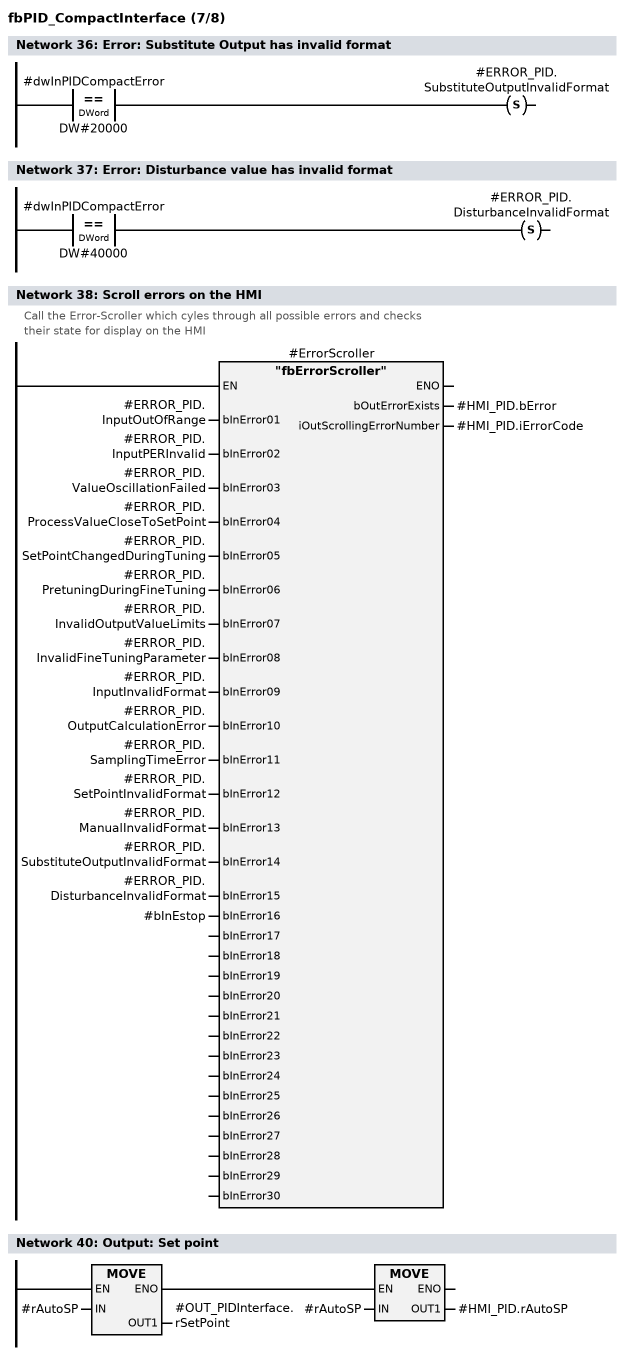
   RUNG wire#powerrail
      { S7_Templates := "SrcType := DWord" } EQ_Contact(in1 := #dwInPIDCompactError, in2 := DW#20000)
      S_Coil( #ERROR_PID.SubstituteOutputInvalidFormat )
   END_RUNG
   // the same network as SCL:
   IF #dwInPIDCompactError = DW#20000 THEN #ERROR_PID.SubstituteOutputInvalidFormat := TRUE; END_IF;
END_REGION

REGION Network 37: Error: Disturbance value has invalid format
   RUNG wire#powerrail
      { S7_Templates := "SrcType := DWord" } EQ_Contact(in1 := #dwInPIDCompactError, in2 := DW#40000)
      S_Coil( #ERROR_PID.DisturbanceInvalidFormat )
   END_RUNG
   // the same network as SCL:
   IF #dwInPIDCompactError = DW#40000 THEN #ERROR_PID.DisturbanceInvalidFormat := TRUE; END_IF;
END_REGION

REGION Network 38: Scroll errors on the HMI
   // Call the Error-Scroller which cyles through all possible errors and checks 
   // their state for display on the HMI
   RUNG wire#powerrail
      #ErrorScroller(bInError01 := #ERROR_PID.InputOutOfRange, bInError02 := #ERROR_PID.InputPERInvalid, bInError03 := #ERROR_PID.ValueOscillationFailed, bInError04 := #ERROR_PID.ProcessValueCloseToSetPoint, bInError05 := #ERROR_PID.SetPointChangedDuringTuning, bInError06 := #ERROR_PID.PretuningDuringFineTuning, bInError07 := #ERROR_PID.InvalidOutputValueLimits, bInError08 := #ERROR_PID.InvalidFineTuningParameter, bInError09 := #ERROR_PID.InputInvalidFormat, bInError10 := #ERROR_PID.OutputCalculationError, bInError11 := #ERROR_PID.SamplingTimeError, bInError12 := #ERROR_PID.SetPointInvalidFormat, bInError13 := #ERROR_PID.ManualInvalidFormat, bInError14 := #ERROR_PID.SubstituteOutputInvalidFormat, bInError15 := #ERROR_PID.DisturbanceInvalidFormat, bInError16 := #bInEstop, bInError17 :=, bInError18 :=, bInError19 :=, bInError20 :=, bInError21 :=, bInError22 :=, bInError23 :=, bInError24 :=, bInError25 :=, bInError26 :=, bInError27 :=, bInError28 :=, bInError29 :=, bInError30 :=, bOutErrorExists => #HMI_PID.bError, iOutScrollingErrorNumber => #HMI_PID.iErrorCode)
   END_RUNG
   // the same network as SCL:
   #ErrorScroller(bInError01 := #ERROR_PID.InputOutOfRange,   // "fbErrorScroller"
                  bInError02 := #ERROR_PID.InputPERInvalid,
                  bInError03 := #ERROR_PID.ValueOscillationFailed,
                  bInError04 := #ERROR_PID.ProcessValueCloseToSetPoint,
                  bInError05 := #ERROR_PID.SetPointChangedDuringTuning,
                  bInError06 := #ERROR_PID.PretuningDuringFineTuning,
                  bInError07 := #ERROR_PID.InvalidOutputValueLimits,
                  bInError08 := #ERROR_PID.InvalidFineTuningParameter,
                  bInError09 := #ERROR_PID.InputInvalidFormat,
                  bInError10 := #ERROR_PID.OutputCalculationError,
                  bInError11 := #ERROR_PID.SamplingTimeError,
                  bInError12 := #ERROR_PID.SetPointInvalidFormat,
                  bInError13 := #ERROR_PID.ManualInvalidFormat,
                  bInError14 := #ERROR_PID.SubstituteOutputInvalidFormat,
                  bInError15 := #ERROR_PID.DisturbanceInvalidFormat,
                  bInError16 := #bInEstop,
                  bOutErrorExists => #HMI_PID.bError,
                  iOutScrollingErrorNumber => #HMI_PID.iErrorCode);
END_REGION

REGION Network 39: --------------------------------------------------------- Outputs ------------------------------------------------------------------
END_REGION

REGION Network 40: Output: Set point
   RUNG wire#powerrail
      Move(in := #rAutoSP, out1 => #OUT_PIDInterface.rSetPoint)
      Move(in := #rAutoSP, out1 => #HMI_PID.rAutoSP)
   END_RUNG
   // the same network as SCL:
   #OUT_PIDInterface.rSetPoint := #rAutoSP;
   #HMI_PID.rAutoSP := #rAutoSP;
END_REGION

REGION Network 41: Output: Process value
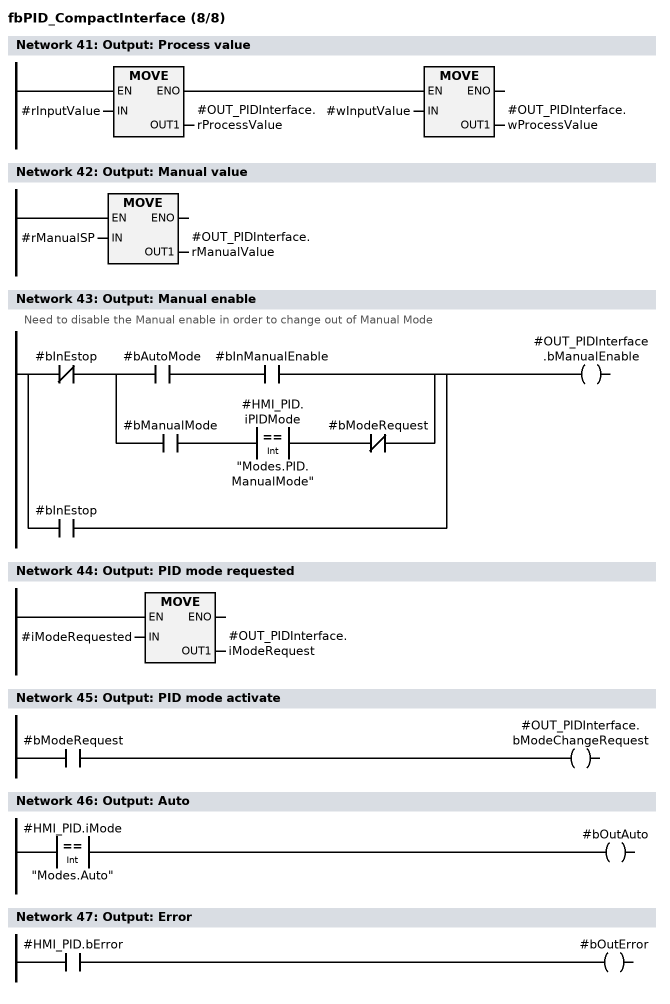
   RUNG wire#powerrail
      Move(in := #rInputValue, out1 => #OUT_PIDInterface.rProcessValue)
      Move(in := #wInputValue, out1 => #OUT_PIDInterface.wProcessValue)
   END_RUNG
   // the same network as SCL:
   #OUT_PIDInterface.rProcessValue := #rInputValue;
   #OUT_PIDInterface.wProcessValue := #wInputValue;
END_REGION

REGION Network 42: Output: Manual value
   RUNG wire#powerrail
      Move(in := #rManualSP, out1 => #OUT_PIDInterface.rManualValue)
   END_RUNG
   // the same network as SCL:
   #OUT_PIDInterface.rManualValue := #rManualSP;
END_REGION

REGION Network 43: Output: Manual enable
   // Need to disable the Manual enable in order to change out of Manual Mode
   RUNG wire#powerrail
      I_Contact( #bInEstop )
      wire#w1
      Contact( #bAutoMode )
      Contact( #bInManualEnable )
      wire#w2
      Coil( #OUT_PIDInterface.bManualEnable )
   END_RUNG
   RUNG wire#w1
      Contact( #bManualMode )
      { S7_Templates := "SrcType := Int" } EQ_Contact(in1 := #HMI_PID.iPIDMode, in2 := "Modes.PID.ManualMode")
      I_Contact( #bModeRequest )
   END_RUNG wire#w2
   RUNG wire#powerrail
      Contact( #bInEstop )
   END_RUNG wire#w2
   // the same network as SCL:
   #OUT_PIDInterface.bManualEnable := (NOT #bInEstop AND ((#bAutoMode AND #bInManualEnable) OR (#bManualMode AND (#HMI_PID.iPIDMode = "Modes.PID.ManualMode") AND NOT #bModeRequest))) OR #bInEstop;
END_REGION

REGION Network 44: Output: PID mode requested
   RUNG wire#powerrail
      Move(in := #iModeRequested, out1 => #OUT_PIDInterface.iModeRequest)
   END_RUNG
   // the same network as SCL:
   #OUT_PIDInterface.iModeRequest := #iModeRequested;
END_REGION

REGION Network 45: Output: PID mode activate
   RUNG wire#powerrail
      Contact( #bModeRequest )
      Coil( #OUT_PIDInterface.bModeChangeRequest )
   END_RUNG
   // the same network as SCL:
   #OUT_PIDInterface.bModeChangeRequest := #bModeRequest;
END_REGION

REGION Network 46: Output: Auto
   RUNG wire#powerrail
      { S7_Templates := "SrcType := Int" } EQ_Contact(in1 := #HMI_PID.iMode, in2 := "Modes.Auto")
      Coil( #bOutAuto )
   END_RUNG
   // the same network as SCL:
   #bOutAuto := #HMI_PID.iMode = "Modes.Auto";
END_REGION

REGION Network 47: Output: Error
   RUNG wire#powerrail
      Contact( #HMI_PID.bError )
      Coil( #bOutError )
   END_RUNG
   // the same network as SCL:
   #bOutError := #HMI_PID.bError;
END_REGION
END_FUNCTION_BLOCK

// folder: Library Blocks/Resources/Communication

FUNCTION_BLOCK "fbAsyncParameterRW_VFD"   // FB125, LAD
TITLE = VFD Acylic Parameter Read and Write
{ S7_Optimized_Access := 'FALSE' }
AUTHOR : JRM
NAME : VFD
VERSION : 0.1
// This block works on Siemens MicroMasters and G120 VFDs
   VAR_TEMP   // added for the SCL form of the ladder/FBD networks
      _w1 : Bool;
   END_VAR
BEGIN

REGION Network 1: ------------------------ Set Values --------------------------
END_REGION

REGION Network 2: Check valid state
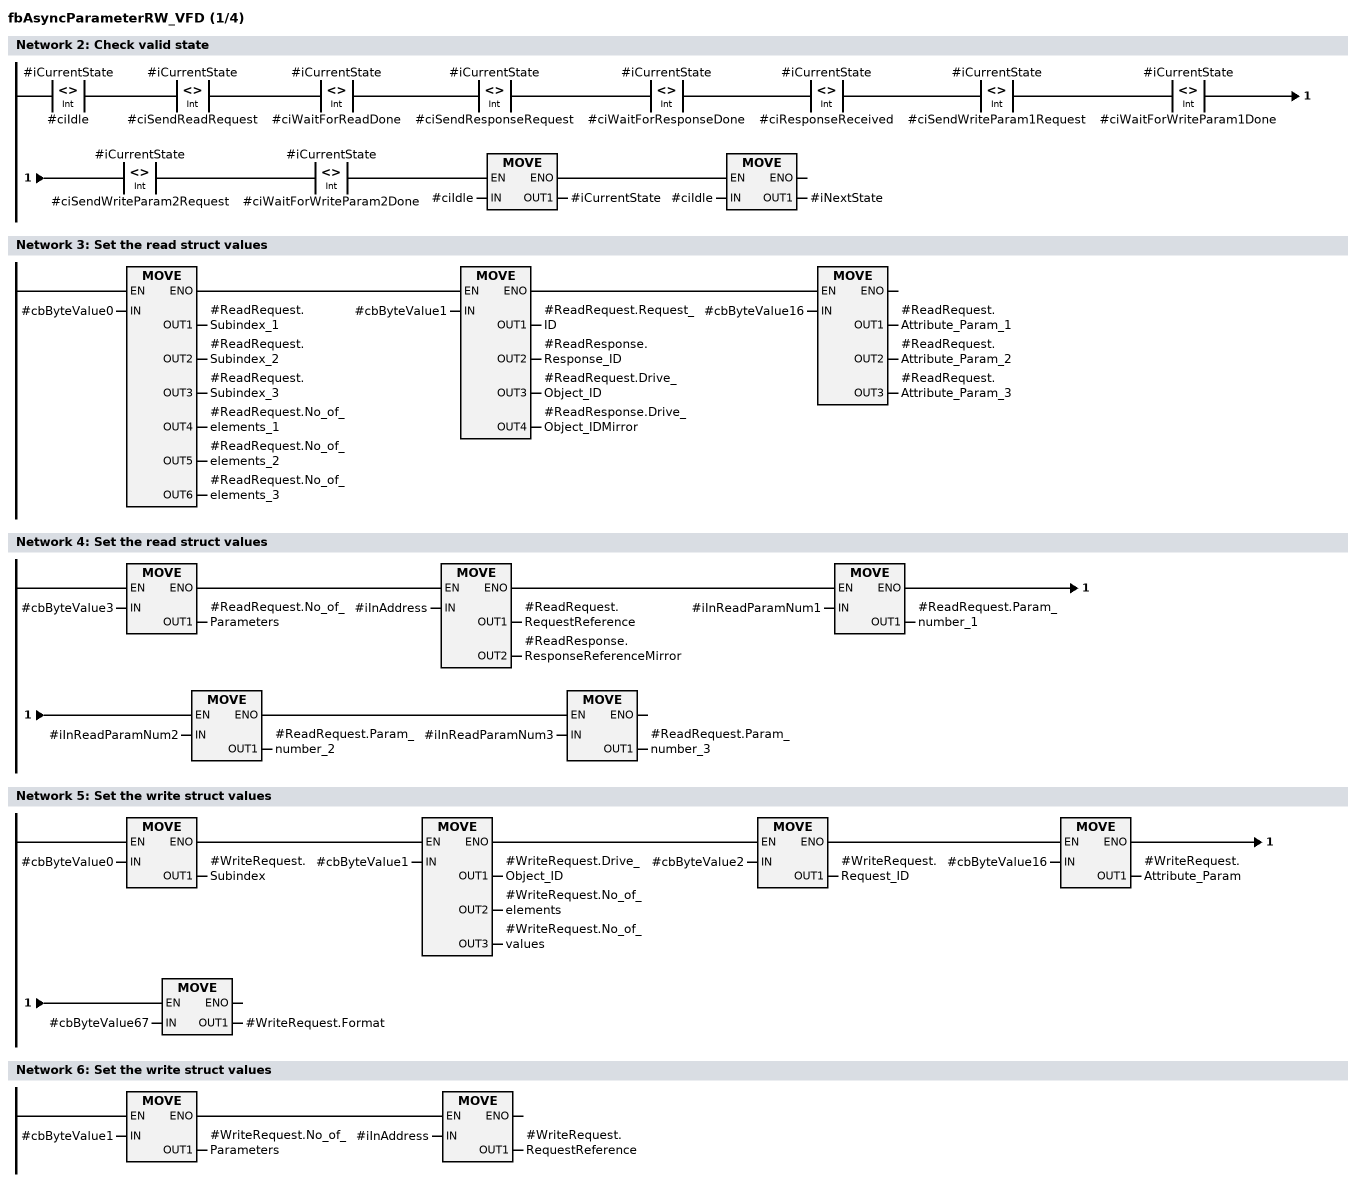
   RUNG wire#powerrail
      { S7_Templates := "SrcType := Int" } NE_Contact(in1 := #iCurrentState, in2 := #ciIdle)
      { S7_Templates := "SrcType := Int" } NE_Contact(in1 := #iCurrentState, in2 := #ciSendReadRequest)
      { S7_Templates := "SrcType := Int" } NE_Contact(in1 := #iCurrentState, in2 := #ciWaitForReadDone)
      { S7_Templates := "SrcType := Int" } NE_Contact(in1 := #iCurrentState, in2 := #ciSendResponseRequest)
      { S7_Templates := "SrcType := Int" } NE_Contact(in1 := #iCurrentState, in2 := #ciWaitForResponseDone)
      { S7_Templates := "SrcType := Int" } NE_Contact(in1 := #iCurrentState, in2 := #ciResponseReceived)
      { S7_Templates := "SrcType := Int" } NE_Contact(in1 := #iCurrentState, in2 := #ciSendWriteParam1Request)
      { S7_Templates := "SrcType := Int" } NE_Contact(in1 := #iCurrentState, in2 := #ciWaitForWriteParam1Done)
      { S7_Templates := "SrcType := Int" } NE_Contact(in1 := #iCurrentState, in2 := #ciSendWriteParam2Request)
      { S7_Templates := "SrcType := Int" } NE_Contact(in1 := #iCurrentState, in2 := #ciWaitForWriteParam2Done)
      { S7_GenerateENO := "TRUE" } Move(in := #ciIdle, out1 => #iCurrentState)
      { S7_GenerateENO := "TRUE" } Move(in := #ciIdle, out1 => #iNextState)
   END_RUNG
   // the same network as SCL:
   // ENO of a box is taken as its EN; it also drops when the box reports an error
   #_w1 := (#iCurrentState <> #ciIdle) AND (#iCurrentState <> #ciSendReadRequest) AND (#iCurrentState <> #ciWaitForReadDone) AND (#iCurrentState <> #ciSendResponseRequest) AND (#iCurrentState <> #ciWaitForResponseDone) AND (#iCurrentState <> #ciResponseReceived) AND (#iCurrentState <> #ciSendWriteParam1Request) AND (#iCurrentState <> #ciWaitForWriteParam1Done) AND (#iCurrentState <> #ciSendWriteParam2Request) AND (#iCurrentState <> #ciWaitForWriteParam2Done);
   IF #_w1 THEN
       #iCurrentState := #ciIdle;
       #iNextState := #ciIdle;
   END_IF;
END_REGION

REGION Network 3: Set the read struct values
   RUNG wire#powerrail
      Move(in := #cbByteValue0, out1 => #ReadRequest.Subindex_1, out2 => #ReadRequest.Subindex_2, out3 => #ReadRequest.Subindex_3, out4 => #ReadRequest.No_of_elements_1, out5 => #ReadRequest.No_of_elements_2, out6 => #ReadRequest.No_of_elements_3)
      Move(in := #cbByteValue1, out1 => #ReadRequest.Request_ID, out2 => #ReadResponse.Response_ID, out3 => #ReadRequest.Drive_Object_ID, out4 => #ReadResponse.Drive_Object_IDMirror)
      { S7_GenerateENO := "TRUE" } Move(in := #cbByteValue16, out1 => #ReadRequest.Attribute_Param_1, out2 => #ReadRequest.Attribute_Param_2, out3 => #ReadRequest.Attribute_Param_3)
   END_RUNG
   // the same network as SCL:
   #ReadRequest.Subindex_1 := #cbByteValue0;
   #ReadRequest.Subindex_2 := #cbByteValue0;
   #ReadRequest.Subindex_3 := #cbByteValue0;
   #ReadRequest.No_of_elements_1 := #cbByteValue0;
   #ReadRequest.No_of_elements_2 := #cbByteValue0;
   #ReadRequest.No_of_elements_3 := #cbByteValue0;
   #ReadRequest.Request_ID := #cbByteValue1;
   #ReadResponse.Response_ID := #cbByteValue1;
   #ReadRequest.Drive_Object_ID := #cbByteValue1;
   #ReadResponse.Drive_Object_IDMirror := #cbByteValue1;
   #ReadRequest.Attribute_Param_1 := #cbByteValue16;
   #ReadRequest.Attribute_Param_2 := #cbByteValue16;
   #ReadRequest.Attribute_Param_3 := #cbByteValue16;
END_REGION

REGION Network 4: Set the read struct values
   RUNG wire#powerrail
      { S7_GenerateENO := "TRUE" } Move(in := #cbByteValue3, out1 => #ReadRequest.No_of_Parameters)
      Move(in := #iInAddress, out1 => #ReadRequest.RequestReference, out2 => #ReadResponse.ResponseReferenceMirror)
      Move(in := #iInReadParamNum1, out1 => #ReadRequest.Param_number_1)
      { S7_GenerateENO := "TRUE" } Move(in := #iInReadParamNum2, out1 => #ReadRequest.Param_number_2)
      { S7_GenerateENO := "TRUE" } Move(in := #iInReadParamNum3, out1 => #ReadRequest.Param_number_3)
   END_RUNG
   // the same network as SCL:
   // ENO of a box is taken as its EN; it also drops when the box reports an error
   #ReadRequest.No_of_Parameters := #cbByteValue3;
   #ReadRequest.RequestReference := #iInAddress;
   #ReadResponse.ResponseReferenceMirror := #iInAddress;
   #ReadRequest.Param_number_1 := #iInReadParamNum1;
   #ReadRequest.Param_number_2 := #iInReadParamNum2;
   #ReadRequest.Param_number_3 := #iInReadParamNum3;
END_REGION

REGION Network 5: Set the write struct values
   RUNG wire#powerrail
      Move(in := #cbByteValue0, out1 => #WriteRequest.Subindex)
      Move(in := #cbByteValue1, out1 => #WriteRequest.Drive_Object_ID, out2 => #WriteRequest.No_of_elements, out3 => #WriteRequest.No_of_values)
      Move(in := #cbByteValue2, out1 => #WriteRequest.Request_ID)
      Move(in := #cbByteValue16, out1 => #WriteRequest.Attribute_Param)
      Move(in := #cbByteValue67, out1 => #WriteRequest.Format)
   END_RUNG
   // the same network as SCL:
   #WriteRequest.Subindex := #cbByteValue0;
   #WriteRequest.Drive_Object_ID := #cbByteValue1;
   #WriteRequest.No_of_elements := #cbByteValue1;
   #WriteRequest.No_of_values := #cbByteValue1;
   #WriteRequest.Request_ID := #cbByteValue2;
   #WriteRequest.Attribute_Param := #cbByteValue16;
   #WriteRequest.Format := #cbByteValue67;
END_REGION

REGION Network 6: Set the write struct values
   RUNG wire#powerrail
      { S7_GenerateENO := "TRUE" } Move(in := #cbByteValue1, out1 => #WriteRequest.No_of_Parameters)
      Move(in := #iInAddress, out1 => #WriteRequest.RequestReference)
   END_RUNG
   // the same network as SCL:
   // ENO of a box is taken as its EN; it also drops when the box reports an error
   #WriteRequest.No_of_Parameters := #cbByteValue1;
   #WriteRequest.RequestReference := #iInAddress;
END_REGION

REGION Network 7: Set the write struct values based on state
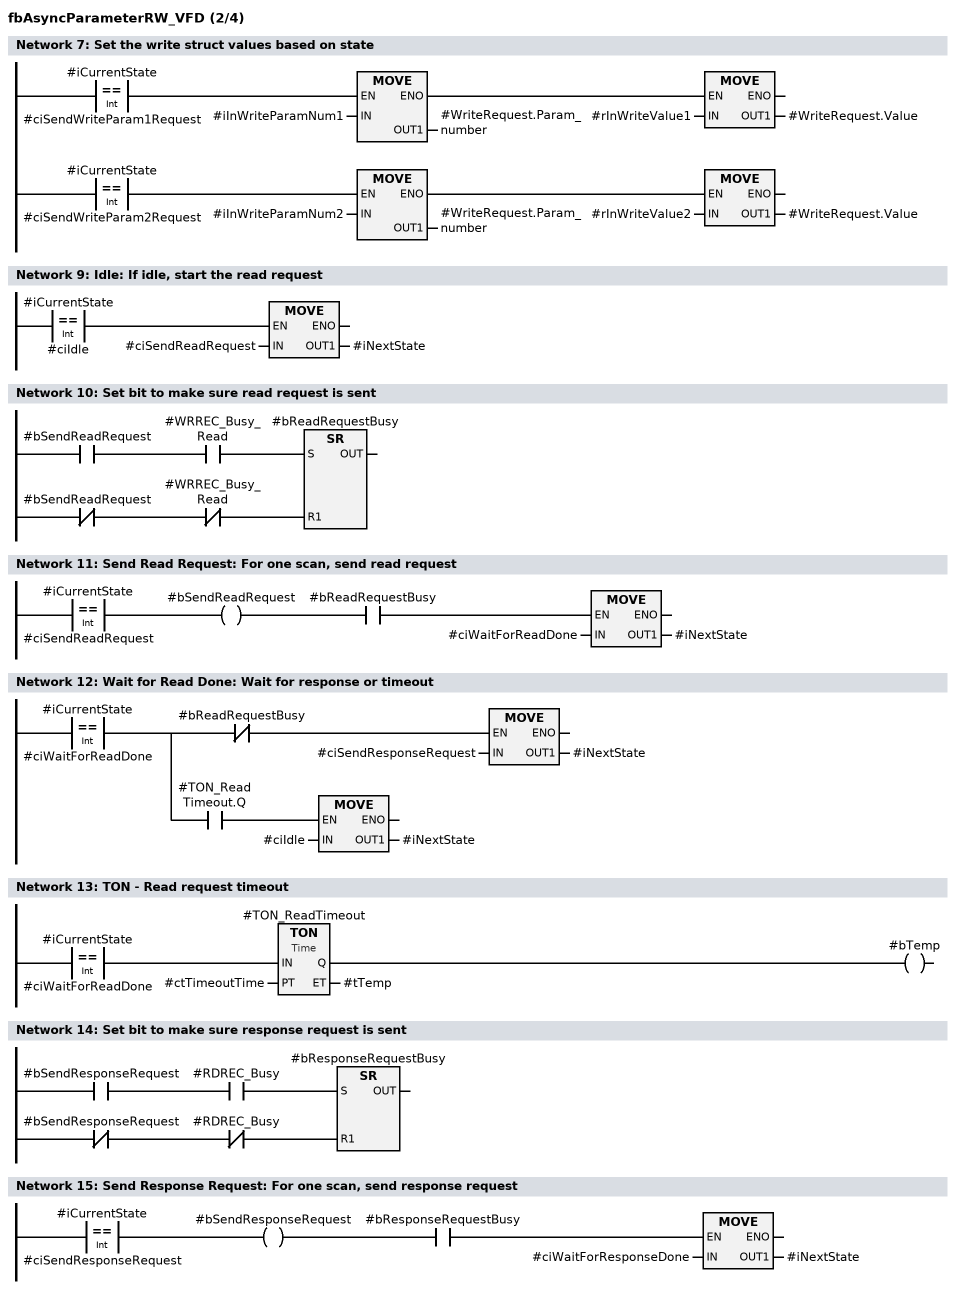
   RUNG wire#powerrail
      { S7_Templates := "SrcType := Int" } EQ_Contact(in1 := #iCurrentState, in2 := #ciSendWriteParam1Request)
      Move(in := #iInWriteParamNum1, out1 => #WriteRequest.Param_number)
      { S7_GenerateENO := "TRUE" } Move(in := #rInWriteValue1, out1 => #WriteRequest.Value)
   END_RUNG
   RUNG wire#powerrail
      { S7_Templates := "SrcType := Int" } EQ_Contact(in1 := #iCurrentState, in2 := #ciSendWriteParam2Request)
      Move(in := #iInWriteParamNum2, out1 => #WriteRequest.Param_number)
      { S7_GenerateENO := "TRUE" } Move(in := #rInWriteValue2, out1 => #WriteRequest.Value)
   END_RUNG
   // the same network as SCL:
   IF #iCurrentState = #ciSendWriteParam1Request THEN
       #WriteRequest.Param_number := #iInWriteParamNum1;
       #WriteRequest.Value := #rInWriteValue1;
   END_IF;
   IF #iCurrentState = #ciSendWriteParam2Request THEN
       #WriteRequest.Param_number := #iInWriteParamNum2;
       #WriteRequest.Value := #rInWriteValue2;
   END_IF;
END_REGION

REGION Network 8: ------------------------ State Logic --------------------------
END_REGION

REGION Network 9: Idle: If idle, start the read request
   RUNG wire#powerrail
      { S7_Templates := "SrcType := Int" } EQ_Contact(in1 := #iCurrentState, in2 := #ciIdle)
      { S7_GenerateENO := "TRUE" } Move(in := #ciSendReadRequest, out1 => #iNextState)
   END_RUNG
   // the same network as SCL:
   IF #iCurrentState = #ciIdle THEN #iNextState := #ciSendReadRequest; END_IF;
END_REGION

REGION Network 10: Set bit to make sure read request is sent
   RUNG wire#powerrail
      Contact( #bSendReadRequest )
      Contact( #WRREC_Busy_Read )
      S_SR(operand := #bReadRequestBusy, r1 := wire#w1)
   END_RUNG
   RUNG wire#powerrail
      I_Contact( #bSendReadRequest )
      I_Contact( #WRREC_Busy_Read )
   END_RUNG wire#w1
   // the same network as SCL:
   IF #bSendReadRequest AND #WRREC_Busy_Read THEN
       #bReadRequestBusy := TRUE;   // SR flip-flop
   END_IF;
   IF NOT #bSendReadRequest AND NOT #WRREC_Busy_Read THEN #bReadRequestBusy := FALSE; END_IF;
END_REGION

REGION Network 11: Send Read Request: For one scan, send read request
   RUNG wire#powerrail
      { S7_Templates := "SrcType := Int" } EQ_Contact(in1 := #iCurrentState, in2 := #ciSendReadRequest)
      Coil( #bSendReadRequest )
      Contact( #bReadRequestBusy )
      Move(in := #ciWaitForReadDone, out1 => #iNextState)
   END_RUNG
   // the same network as SCL:
   #bSendReadRequest := #iCurrentState = #ciSendReadRequest;
   IF #bSendReadRequest AND #bReadRequestBusy THEN #iNextState := #ciWaitForReadDone; END_IF;
END_REGION

REGION Network 12: Wait for Read Done: Wait for response or timeout
   RUNG wire#powerrail
      { S7_Templates := "SrcType := Int" } EQ_Contact(in1 := #iCurrentState, in2 := #ciWaitForReadDone)
      wire#w1
      I_Contact( #bReadRequestBusy )
      { S7_GenerateENO := "TRUE" } Move(in := #ciSendResponseRequest, out1 => #iNextState)
   END_RUNG
   RUNG wire#w1
      Contact( #TON_ReadTimeout.Q )
      { S7_GenerateENO := "TRUE" } Move(in := #ciIdle, out1 => #iNextState)
   END_RUNG
   // the same network as SCL:
   #_w1 := #iCurrentState = #ciWaitForReadDone;
   IF #_w1 AND NOT #bReadRequestBusy THEN #iNextState := #ciSendResponseRequest; END_IF;
   IF #_w1 AND #TON_ReadTimeout.Q THEN #iNextState := #ciIdle; END_IF;
END_REGION

REGION Network 13: TON - Read request timeout
   #TON_ReadTimeout.TON(IN := #iCurrentState = #ciWaitForReadDone, PT := #ctTimeoutTime, ET => #tTemp);
   #bTemp := #TON_ReadTimeout.Q;
END_REGION

REGION Network 14: Set bit to make sure response request is sent
   RUNG wire#powerrail
      Contact( #bSendResponseRequest )
      Contact( #RDREC_Busy )
      S_SR(operand := #bResponseRequestBusy, r1 := wire#w1)
   END_RUNG
   RUNG wire#powerrail
      I_Contact( #bSendResponseRequest )
      I_Contact( #RDREC_Busy )
   END_RUNG wire#w1
   // the same network as SCL:
   IF #bSendResponseRequest AND #RDREC_Busy THEN
       #bResponseRequestBusy := TRUE;   // SR flip-flop
   END_IF;
   IF NOT #bSendResponseRequest AND NOT #RDREC_Busy THEN #bResponseRequestBusy := FALSE; END_IF;
END_REGION

REGION Network 15: Send Response Request: For one scan, send response request
   RUNG wire#powerrail
      { S7_Templates := "SrcType := Int" } EQ_Contact(in1 := #iCurrentState, in2 := #ciSendResponseRequest)
      Coil( #bSendResponseRequest )
      Contact( #bResponseRequestBusy )
      Move(in := #ciWaitForResponseDone, out1 => #iNextState)
   END_RUNG
   // the same network as SCL:
   #bSendResponseRequest := #iCurrentState = #ciSendResponseRequest;
   IF #bSendResponseRequest AND #bResponseRequestBusy THEN #iNextState := #ciWaitForResponseDone; END_IF;
END_REGION

REGION Network 16: Wait for Resonse Done: Wait for response or timeout
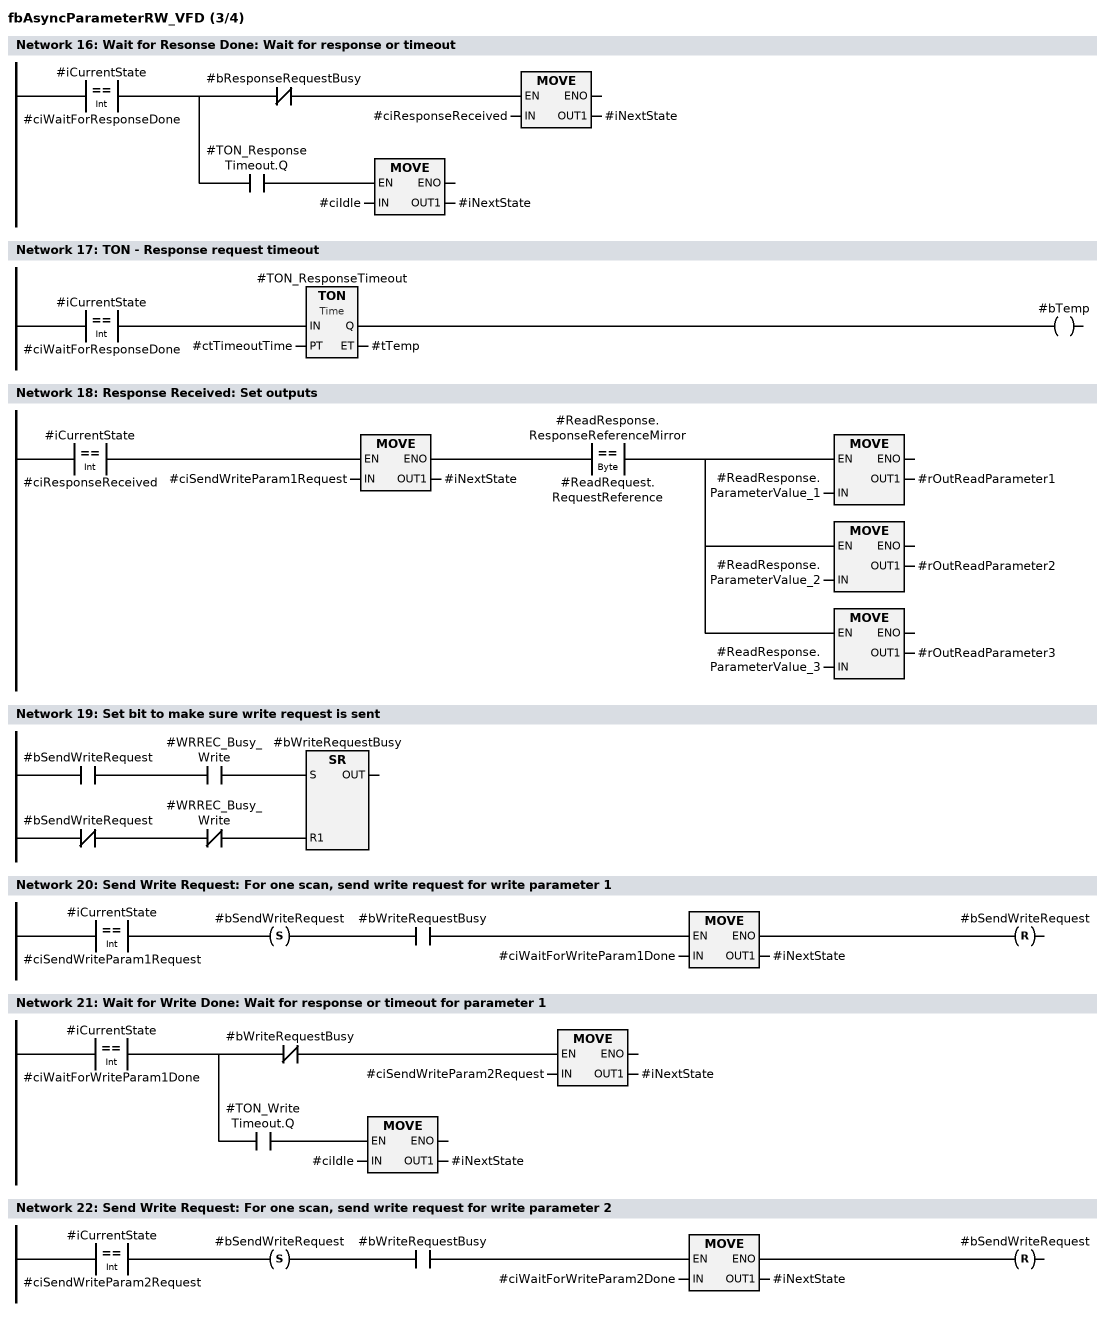
   RUNG wire#powerrail
      { S7_Templates := "SrcType := Int" } EQ_Contact(in1 := #iCurrentState, in2 := #ciWaitForResponseDone)
      wire#w1
      I_Contact( #bResponseRequestBusy )
      { S7_GenerateENO := "TRUE" } Move(in := #ciResponseReceived, out1 => #iNextState)
   END_RUNG
   RUNG wire#w1
      Contact( #TON_ResponseTimeout.Q )
      { S7_GenerateENO := "TRUE" } Move(in := #ciIdle, out1 => #iNextState)
   END_RUNG
   // the same network as SCL:
   #_w1 := #iCurrentState = #ciWaitForResponseDone;
   IF #_w1 AND NOT #bResponseRequestBusy THEN #iNextState := #ciResponseReceived; END_IF;
   IF #_w1 AND #TON_ResponseTimeout.Q THEN #iNextState := #ciIdle; END_IF;
END_REGION

REGION Network 17: TON - Response request timeout
   #TON_ResponseTimeout.TON(IN := #iCurrentState = #ciWaitForResponseDone, PT := #ctTimeoutTime, ET => #tTemp);
   #bTemp := #TON_ResponseTimeout.Q;
END_REGION

REGION Network 18: Response Received: Set outputs
   RUNG wire#powerrail
      { S7_Templates := "SrcType := Int" } EQ_Contact(in1 := #iCurrentState, in2 := #ciResponseReceived)
      { S7_GenerateENO := "TRUE" } Move(in := #ciSendWriteParam1Request, out1 => #iNextState)
      { S7_Templates := "SrcType := Byte" } EQ_Contact(in1 := #ReadResponse.ResponseReferenceMirror, in2 := #ReadRequest.RequestReference)
      wire#w1
      { S7_GenerateENO := "TRUE" } Move(in := #ReadResponse.ParameterValue_1, out1 => #rOutReadParameter1)
   END_RUNG
   RUNG wire#w1
      { S7_GenerateENO := "TRUE" } Move(in := #ReadResponse.ParameterValue_2, out1 => #rOutReadParameter2)
   END_RUNG
   RUNG wire#w1
      { S7_GenerateENO := "TRUE" } Move(in := #ReadResponse.ParameterValue_3, out1 => #rOutReadParameter3)
   END_RUNG
   // the same network as SCL:
   // ENO of a box is taken as its EN; it also drops when the box reports an error
   #_w1 := #iCurrentState = #ciResponseReceived;
   IF #_w1 THEN #iNextState := #ciSendWriteParam1Request; END_IF;
   IF #_w1 AND (#ReadResponse.ResponseReferenceMirror = #ReadRequest.RequestReference) THEN
       #rOutReadParameter1 := #ReadResponse.ParameterValue_1;
       #rOutReadParameter2 := #ReadResponse.ParameterValue_2;
       #rOutReadParameter3 := #ReadResponse.ParameterValue_3;
   END_IF;
END_REGION

REGION Network 19: Set bit to make sure write request is sent
   RUNG wire#powerrail
      Contact( #bSendWriteRequest )
      Contact( #WRREC_Busy_Write )
      S_SR(operand := #bWriteRequestBusy, r1 := wire#w1)
   END_RUNG
   RUNG wire#powerrail
      I_Contact( #bSendWriteRequest )
      I_Contact( #WRREC_Busy_Write )
   END_RUNG wire#w1
   // the same network as SCL:
   IF #bSendWriteRequest AND #WRREC_Busy_Write THEN
       #bWriteRequestBusy := TRUE;   // SR flip-flop
   END_IF;
   IF NOT #bSendWriteRequest AND NOT #WRREC_Busy_Write THEN #bWriteRequestBusy := FALSE; END_IF;
END_REGION

REGION Network 20: Send Write Request: For one scan, send write request for write parameter 1
   RUNG wire#powerrail
      { S7_Templates := "SrcType := Int" } EQ_Contact(in1 := #iCurrentState, in2 := #ciSendWriteParam1Request)
      S_Coil( #bSendWriteRequest )
      Contact( #bWriteRequestBusy )
      Move(in := #ciWaitForWriteParam1Done, out1 => #iNextState)
      R_Coil( #bSendWriteRequest )
   END_RUNG
   // the same network as SCL:
   #_w1 := #iCurrentState = #ciSendWriteParam1Request;
   IF #_w1 THEN #bSendWriteRequest := TRUE; END_IF;
   IF #_w1 AND #bWriteRequestBusy THEN
       #iNextState := #ciWaitForWriteParam1Done;
       #bSendWriteRequest := FALSE;
   END_IF;
END_REGION

REGION Network 21: Wait for Write Done: Wait for response or timeout for parameter 1
   RUNG wire#powerrail
      { S7_Templates := "SrcType := Int" } EQ_Contact(in1 := #iCurrentState, in2 := #ciWaitForWriteParam1Done)
      wire#w1
      I_Contact( #bWriteRequestBusy )
      { S7_GenerateENO := "TRUE" } Move(in := #ciSendWriteParam2Request, out1 => #iNextState)
   END_RUNG
   RUNG wire#w1
      Contact( #TON_WriteTimeout.Q )
      { S7_GenerateENO := "TRUE" } Move(in := #ciIdle, out1 => #iNextState)
   END_RUNG
   // the same network as SCL:
   #_w1 := #iCurrentState = #ciWaitForWriteParam1Done;
   IF #_w1 AND NOT #bWriteRequestBusy THEN #iNextState := #ciSendWriteParam2Request; END_IF;
   IF #_w1 AND #TON_WriteTimeout.Q THEN #iNextState := #ciIdle; END_IF;
END_REGION

REGION Network 22: Send Write Request: For one scan, send write request for write parameter 2
   RUNG wire#powerrail
      { S7_Templates := "SrcType := Int" } EQ_Contact(in1 := #iCurrentState, in2 := #ciSendWriteParam2Request)
      S_Coil( #bSendWriteRequest )
      Contact( #bWriteRequestBusy )
      Move(in := #ciWaitForWriteParam2Done, out1 => #iNextState)
      R_Coil( #bSendWriteRequest )
   END_RUNG
   // the same network as SCL:
   #_w1 := #iCurrentState = #ciSendWriteParam2Request;
   IF #_w1 THEN #bSendWriteRequest := TRUE; END_IF;
   IF #_w1 AND #bWriteRequestBusy THEN
       #iNextState := #ciWaitForWriteParam2Done;
       #bSendWriteRequest := FALSE;
   END_IF;
END_REGION

REGION Network 23: Wait for Write Done: Wait for response or timeout for parameter 2
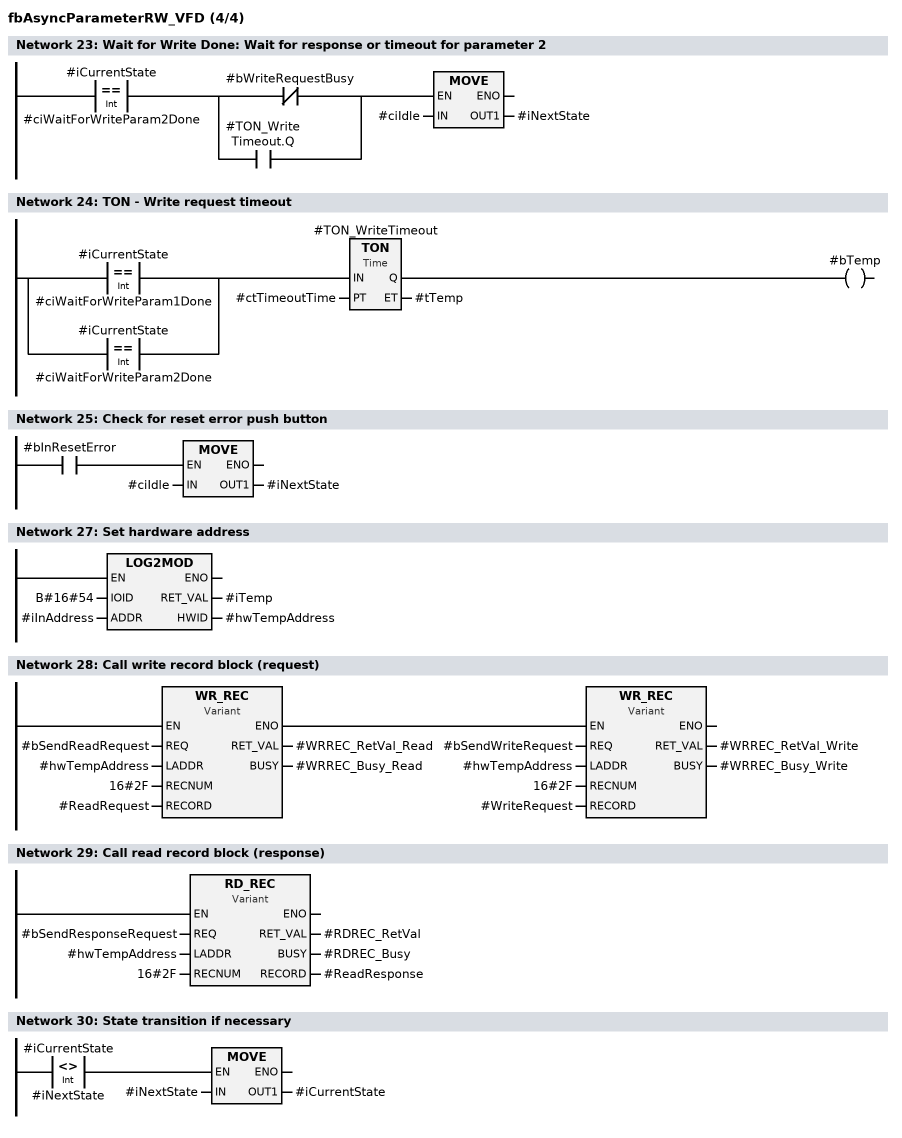
   RUNG wire#powerrail
      { S7_Templates := "SrcType := Int" } EQ_Contact(in1 := #iCurrentState, in2 := #ciWaitForWriteParam2Done)
      wire#w1
      I_Contact( #bWriteRequestBusy )
      wire#w2
      { S7_GenerateENO := "TRUE" } Move(in := #ciIdle, out1 => #iNextState)
   END_RUNG
   RUNG wire#w1
      Contact( #TON_WriteTimeout.Q )
   END_RUNG wire#w2
   // the same network as SCL:
   IF (#iCurrentState = #ciWaitForWriteParam2Done) AND (NOT #bWriteRequestBusy OR #TON_WriteTimeout.Q) THEN
       #iNextState := #ciIdle;
   END_IF;
END_REGION

REGION Network 24: TON - Write request timeout
   #TON_WriteTimeout.TON(IN := (#iCurrentState = #ciWaitForWriteParam1Done) OR (#iCurrentState = #ciWaitForWriteParam2Done),
                         PT := #ctTimeoutTime,
                         ET => #tTemp);
   #bTemp := #TON_WriteTimeout.Q;
END_REGION

REGION Network 25: Check for reset error push button
   RUNG wire#powerrail
      Contact( #bInResetError )
      Move(in := #ciIdle, out1 => #iNextState)
   END_RUNG
   // the same network as SCL:
   IF #bInResetError THEN #iNextState := #ciIdle; END_IF;
END_REGION

REGION Network 26: --------------------- Call Read Blocks ---------------------
END_REGION

REGION Network 27: Set hardware address
   #iTemp := LOG2MOD(IOID := B#16#54, ADDR := #iInAddress, HWID => #hwTempAddress);
END_REGION

REGION Network 28: Call write record block (request)
   // ENO of a box is taken as its EN; it also drops when the box reports an error
   #WRREC_RetVal_Read := WR_REC(REQ := #bSendReadRequest,
                           LADDR := #hwTempAddress,
                           RECNUM := 16#2F,
                           RECORD := #ReadRequest,
                           BUSY => #WRREC_Busy_Read);
   #WRREC_RetVal_Write := WR_REC(REQ := #bSendWriteRequest,
                           LADDR := #hwTempAddress,
                           RECNUM := 16#2F,
                           RECORD := #WriteRequest,
                           BUSY => #WRREC_Busy_Write);
END_REGION

REGION Network 29: Call read record block (response)
   #RDREC_RetVal := RD_REC(REQ := #bSendResponseRequest,
                           LADDR := #hwTempAddress,
                           RECNUM := 16#2F,
                           BUSY => #RDREC_Busy,
                           RECORD => #ReadResponse);
END_REGION

REGION Network 30: State transition if necessary
   RUNG wire#powerrail
      { S7_Templates := "SrcType := Int" } NE_Contact(in1 := #iCurrentState, in2 := #iNextState)
      { S7_GenerateENO := "TRUE" } Move(in := #iNextState, out1 => #iCurrentState)
   END_RUNG
   // the same network as SCL:
   IF #iCurrentState <> #iNextState THEN #iCurrentState := #iNextState; END_IF;
END_REGION
END_FUNCTION_BLOCK

// folder: Library Blocks/Resources/Conversion

FUNCTION "fcSwapBytes" : Void   // FC300, LAD
TITLE = Swap the bytes in a word
{ S7_Optimized_Access := 'FALSE' }
AUTHOR : DMC
FAMILY : LowLevel
VERSION : 0.1
// High byte and Low Byte are swapped
BEGIN

REGION Network 1: Swap the bytes
   // High byte and Low Byte are swapped
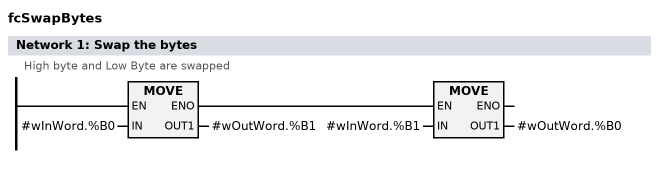
   RUNG wire#powerrail
      { S7_GenerateENO := "TRUE" } Move(in := #wInWord.%B0, out1 => #wOutWord.%B1)
      { S7_GenerateENO := "TRUE" } Move(in := #wInWord.%B1, out1 => #wOutWord.%B0)
   END_RUNG
   // the same network as SCL:
   // ENO of a box is taken as its EN; it also drops when the box reports an error
   #wOutWord.%B1 := #wInWord.%B0;
   #wOutWord.%B0 := #wInWord.%B1;
END_REGION
END_FUNCTION

FUNCTION "fcWordToBits" : Void   // FC1000, LAD
TITLE = Breaks A Word Into Individual Bits
{ S7_Optimized_Access := 'FALSE' }
AUTHOR : DMC
FAMILY : LowLevel
VERSION : 0.1
BEGIN

REGION Network 1: Bit0
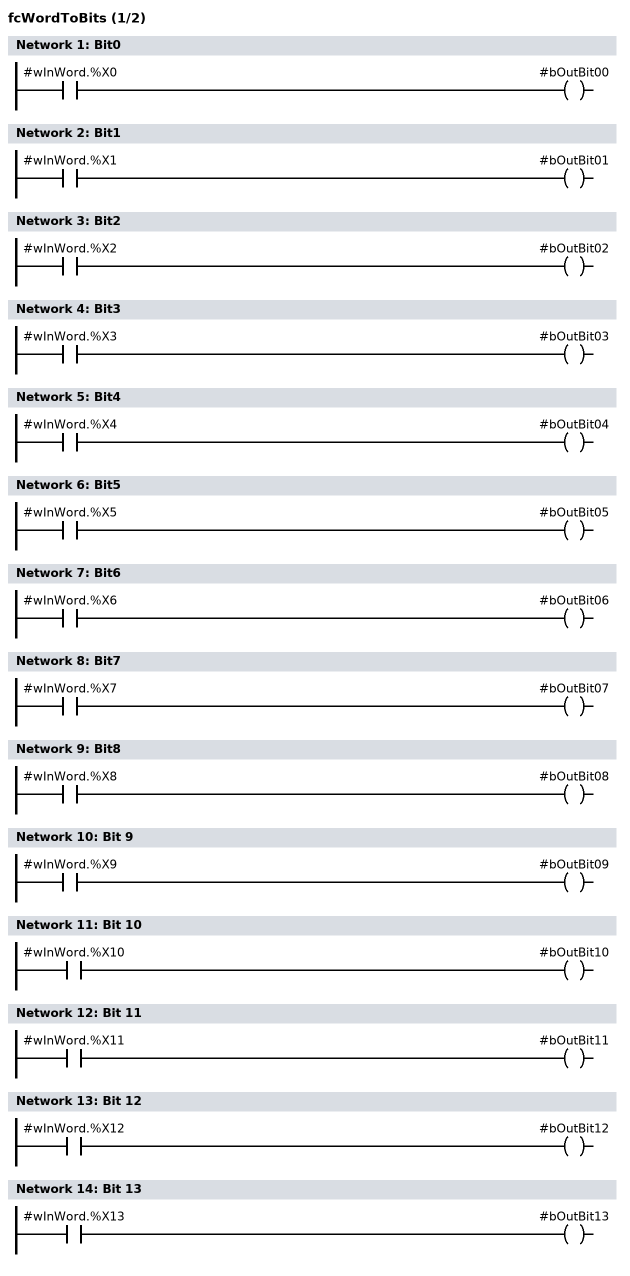
   RUNG wire#powerrail
      Contact( #wInWord.%X0 )
      Coil( #bOutBit00 )
   END_RUNG
   // the same network as SCL:
   #bOutBit00 := #wInWord.%X0;
END_REGION

REGION Network 2: Bit1
   RUNG wire#powerrail
      Contact( #wInWord.%X1 )
      Coil( #bOutBit01 )
   END_RUNG
   // the same network as SCL:
   #bOutBit01 := #wInWord.%X1;
END_REGION

REGION Network 3: Bit2
   RUNG wire#powerrail
      Contact( #wInWord.%X2 )
      Coil( #bOutBit02 )
   END_RUNG
   // the same network as SCL:
   #bOutBit02 := #wInWord.%X2;
END_REGION

REGION Network 4: Bit3
   RUNG wire#powerrail
      Contact( #wInWord.%X3 )
      Coil( #bOutBit03 )
   END_RUNG
   // the same network as SCL:
   #bOutBit03 := #wInWord.%X3;
END_REGION

REGION Network 5: Bit4
   RUNG wire#powerrail
      Contact( #wInWord.%X4 )
      Coil( #bOutBit04 )
   END_RUNG
   // the same network as SCL:
   #bOutBit04 := #wInWord.%X4;
END_REGION

REGION Network 6: Bit5
   RUNG wire#powerrail
      Contact( #wInWord.%X5 )
      Coil( #bOutBit05 )
   END_RUNG
   // the same network as SCL:
   #bOutBit05 := #wInWord.%X5;
END_REGION

REGION Network 7: Bit6
   RUNG wire#powerrail
      Contact( #wInWord.%X6 )
      Coil( #bOutBit06 )
   END_RUNG
   // the same network as SCL:
   #bOutBit06 := #wInWord.%X6;
END_REGION

REGION Network 8: Bit7
   RUNG wire#powerrail
      Contact( #wInWord.%X7 )
      Coil( #bOutBit07 )
   END_RUNG
   // the same network as SCL:
   #bOutBit07 := #wInWord.%X7;
END_REGION

REGION Network 9: Bit8
   RUNG wire#powerrail
      Contact( #wInWord.%X8 )
      Coil( #bOutBit08 )
   END_RUNG
   // the same network as SCL:
   #bOutBit08 := #wInWord.%X8;
END_REGION
